(* CODESYS project JSON Utilities SL Example.project
   Title: JSON Utilities SL Example
   Author: CODESYS Development GmbH
   Company: CODESYS

Project tree, tasks and I/O mapping:
  Device : CODESYS Control for Raspberry Pi 64 SL, CODESYS, order no. 2302000009, version 4.18.0.0
    application JSONFindValueExample
      libraries: Standard, 3.5.18.0 (System); VisuDialogs, * (System); CAA FB Factory, * (CAA Technical Workgroup); JSON Utilities SL, 1.11.0.0 (CODESYS)
      task MainTask (cyclic, interval t#20ms, priority 1) calls PLC_PRG
      task VISU_TASK (cyclic, interval 100 ms, priority 31) calls VisuElems.Visu_Prg
      program PLC_PRG [CFC]
      visualisation Visualization
      image pool ImagePool
    application JSONFileExample
      libraries: Standard, 3.5.18.0 (System); VisuDialogs, * (System); CAA FB Factory, * (CAA Technical Workgroup); JSON Utilities SL, 1.11.0.0 (CODESYS)
      task MainTask (cyclic, interval t#20ms, priority 1) calls PLC_PRG
      task VISU_TASK (cyclic, interval 100 ms, priority 31) calls VisuElems.Visu_Prg
      program PLC_PRG [CFC]
      visualisation Visualization
      image pool ImagePool
    application JSONArrayExample
      libraries: Standard, 3.5.18.0 (System); VisuDialogs, * (System); CAA FB Factory, * (CAA Technical Workgroup); JSON Utilities SL, 1.11.0.0 (CODESYS)
      task MainTask (cyclic, interval t#20ms, priority 1) calls PLC_PRG
      task VISU_TASK (cyclic, interval 100 ms, priority 31) calls VisuElems.Visu_Prg
      program PLC_PRG [CFC]
      visualisation Visualization
      image pool ImagePool
    application JSONDataExample
      libraries: CAA FB Factory, * (CAA Technical Workgroup); JSON Utilities SL, 1.11.0.0 (CODESYS)
      task Task (cyclic, interval t#20ms, priority 1) calls PLC_PRG
      program PLC_PRG [ST]
    SoftMotion General Axis Pool
    GPIOs_A_B : GPIOs A/B, CODESYS, version 4.18.0.0
        unmapped channels: digital inputs (GPIO0..GPIO31), digital outputs (GPIO0..GPIO31)
    Onewire
    Camera device
      <Empty>
    SPI
    I²C
  text list GlobalTextList
  function block Element2StringArray [ST]
  5ce3da45-db07-42e7-a21c-a00fff4ed8f6|C:\Users\a.werner\Documents\background.jpg
  5ce3da45-db07-42e7-a21c-a00fff4ed8f6|C:\Users\a.werner\Documents\background.jpg
  5ce3da45-db07-42e7-a21c-a00fff4ed8f6|C:\Users\a.werner\Documents\background.jpg
*)

// Device/JSONFindValueExample/PLC_PRG
// This program loads the demo file 'test.json' and finds the value of the first key in the file. 
PROGRAM PLC_PRG
VAR
	sFileName : STRING(255) := 'res/test.json';	

	jsonDataFactory : JSON.JSONDataFactory;
	eDataFactoryError : FBF.ERROR; // Error code: 0: OK, 30103: no more memory 
	pJSONData : POINTER TO JSON.JSONData := jsonDataFactory.Create(eError => eDataFactoryError);

	JSONFileReader_0: JSON.JSONFileReader;
	xStart : BOOL;
	xFindValue : BOOL;
	wsKey : WSTRING := "Vorname";
	element : JSON.JSONElement;
	FindFirstValueByKey_0: JSON.FindFirstValueByKey;
	wsValue: WSTRING(JSON.GParams.g_diMaxStringSize);
END_VAR

// Load the example file 'c:\temp\test.json'
JSONFileReader_0(xExecute := xStart, sFileName := sFileName, jsonData := pJSONData^); // JSON.JSONFileReader
// Find a value by key
FindFirstValueByKey_0(xExecute := xFindValue, wsKey := wsKey, diStartIndex := 0, jsonData := pJSONData^); // JSON.FindFirstValueByKey
JSON.JSONElementToString(element := FindFirstValueByKey_0.jsonElement, wsResult := wsValue);

END_PROGRAM

// Device/JSONFileExample/PLC_PRG
// This program shows how to read and write JSON files.
PROGRAM PLC_PRG
VAR
	// JSON data container
	jsonDataFactory : JSON.JSONDataFactory; // Factory to create a JSONData function block. 
	eDataFactoryError : FBF.ERROR; // Error code: 0: OK, 30103: no more memory
	pJSONData : POINTER TO JSON.JSONData := jsonDataFactory.Create(eError => eDataFactoryError); // Result of Create is a pointer to JSONData
	
	// Reader
	JSONFileReader_0: JSON.JSONFileReader; 
	wsFilenameRead : STRING(255) := 'res/test.json';
	xReadFile : BOOL;
	
	// Writer
	JSONFileWriter_0: JSON.JSONFileWriter;
	wsFilenameWrite : STRING(255) := 'res/testWrite.json';
	xWriteFile : BOOL;
	
	// Helper array for visu
	awsData :  ARRAY[0..3, 0..500] OF WSTRING(JSON.GParams.g_diMaxStringSize);
	element2StringArray : Element2StringArray; // Function block to convert the sample data into an array of WSTRINGs (only for visualization)
END_VAR

// Convert the result into an array of WSTRINGs (only for visualization)
element2StringArray(xExecute := JSONFileReader_0.xDone, jsonData := pJSONData^, awsDataArray := awsData);
// Load the example file 'c:\temp\test.json'
JSONFileReader_0(xExecute := xReadFile, sFileName := wsFilenameRead, jsonData := pJSONData^); // JSON.JSONFileReader
// Write a JSON file
JSONFileWriter_0(
    xExecute := xWriteFile,
    sFileName := wsFilenameWrite,
    eEncoding := JSON.Encoding.UTF_8,
    jsonData := pJSONData^); // JSON.JSONFileWriter

END_PROGRAM

// Element2StringArray
// Helper function to convert the JSON elements to an array of WSTRINGs.
FUNCTION_BLOCK Element2StringArray
VAR_INPUT
	xExecute : BOOL; // Starts converting..
END_VAR
VAR_IN_OUT
	jsonData : JSON.JSONData;
	awsDataArray : ARRAY[0..3, 0..500] OF WSTRING(JSON.GParams.g_diMaxStringSize);
END_VAR
VAR
	diCounter : DINT;
	irow, icol : INT;
	element : JSON.JSONElement;
	j, i : INT;
END_VAR

IF xExecute = FALSE THEN
	RETURN;
END_IF
diCounter := 0;
irow := 0;
WHILE irow < 500 AND diCounter < JSON.GParams.g_diMaxElements DO
	jsonData.GetElementByIndex(diIndex := diCounter, jsonElement => element);
	IF element.eType = JSON.JSONType.NONE THEN
		FOR j := irow TO 500 DO
			FOR i := 0 TO 3 DO
				awsDataArray[i, j] := "";
			END_FOR	
		END_FOR
		RETURN;
	END_IF
	icol := 0;	
	
	// Index
	awsDataArray[icol, irow] := DINT_TO_WSTRING(element.diIndex);
	icol := icol + 1;
	
	// Parent Index
	awsDataArray[icol, irow] := DINT_TO_WSTRING(element.diParentIndex);
	icol := icol + 1;
	
	// Type
	IF element.eType = JSON.JSONType.BOOL_VALUE THEN
		awsDataArray[icol, irow] := "Bool";
	ELSIF element.eType = JSON.JSONType.LINT_VALUE THEN
		awsDataArray[icol, irow] := "LInt";
	ELSIF element.eType = JSON.JSONType.JSON_ARRAY THEN
		awsDataArray[icol, irow] := "Array";
	ELSIF element.eType = JSON.JSONType.JSON_OBJECT THEN
		awsDataArray[icol, irow] := "Object";
	ELSIF element.eType = JSON.JSONType.KEY THEN
		awsDataArray[icol, irow] := "Key";
	ELSIF element.eType = JSON.JSONType.NONE THEN
		awsDataArray[icol, irow] := "None";
	ELSIF element.eType = JSON.JSONType.NULL THEN
		awsDataArray[icol, irow] := "Null";
	ELSIF element.eType = JSON.JSONType.LREAL_VALUE THEN
		awsDataArray[icol, irow] := "LReal";
	ELSIF element.eType = JSON.JSONType.WSTRING_VALUE THEN
		awsDataArray[icol, irow] := "String";
	ELSE
		awsDataArray[icol, irow] := "Unknown";
	END_IF	
	icol := icol + 1;
	
	// Value
	IF element.eType = JSON.JSONType.BOOL_VALUE THEN
		awsDataArray[icol, irow] := BOOL_TO_WSTRING(element.value.xValue);
	ELSIF element.eType = JSON.JSONType.LINT_VALUE THEN
		awsDataArray[icol, irow] := LINT_TO_WSTRING(element.value.liValue);
	ELSIF element.eType = JSON.JSONType.KEY OR element.eType = JSON.JSONType.WSTRING_VALUE THEN
		awsDataArray[icol, irow] := element.value.wsValue;
	ELSIF element.eType = JSON.JSONType.LREAL_VALUE THEN
		awsDataArray[icol, irow] := LREAL_TO_WSTRING(element.value.lrValue);	
	ELSIF element.eType = JSON.JSONType.NULL THEN
		awsDataArray[icol, irow] := "Null";	
	ELSE
		awsDataArray[icol, irow] := "";	
	END_IF
	irow := irow + 1;
	diCounter := diCounter + 1;	
END_WHILE

END_FUNCTION_BLOCK

// Device/JSONArrayExample/PLC_PRG
// This program shows how to read and write JSON arrays.
PROGRAM PLC_PRG
VAR
	// JSON data container
	jsonDataFactory : JSON.JSONDataFactory; // Factory to create a JSONData function block. 
	eDataFactoryError : FBF.ERROR; // Error code: 0: OK, 30103: no more memory
	pJSONData : POINTER TO JSON.JSONData := jsonDataFactory.Create(eError => eDataFactoryError); // Result of Create is a pointer to JSONData
	
	// Reader
	JSONByteArrayReader_0: JSON.JSONByteArrayReader;	
	xRead : BOOL;
	// Demo data
	wsData : WSTRING(1024) := "{
  $0022Herausgeber$0022: $0022Xema$0022,
  $0022Nummer$0022: $00221234-5678-9012-3456$0022,
  $0022Deckung$0022: -0.444,
  $0022Waehrung$0022: $0022EURO$0022,
  $0022Inhaber$0022: 
  {
    $0022Name$0022: $0022Mustermann$0022,
    $0022Vorname$0022: $0022Max$0022,
    $0022maennlich$0022: true,
    $0022Hobbys$0022: [ $0022Reiten$0022, $0022Golfen$0022, $0022Lesen$0022 ],
    $0022Alter$0022: 42,
    $0022Kinder$0022: [],
    $0022Partner$0022: null
  }
}";
	
	// Writer
	JSONByteArrayWriter_0: JSON.JSONByteArrayWriter;
	wsWriteData : WSTRING(1024) := ""; // The result of the Writer
	xWrite : BOOL;
	
	// Helper array for visu
	awsData :  ARRAY[0..3, 0..500] OF WSTRING(JSON.GParams.g_diMaxStringSize);	
	element2StringArray : Element2StringArray; // Function block to convert the sample data into an array of WSTRINGs (only for visualization)
END_VAR

// Read JSON data from WSTRING
JSONByteArrayReader_0(xExecute := xRead, pwData := ADR(wsData), jsonData := pJSONData^); // JSON.JSONByteArrayReader
// Convert the result into an array of WSTRINGs (only for visualization)
element2StringArray(xExecute := JSONByteArrayReader_0.xDone, jsonData := pJSONData^, awsDataArray := awsData);
// Read JSON data to WSTRING
JSONByteArrayWriter_0(
    xExecute := xWrite,
    pwData := ADR(wsWriteData),
    udiSize := SIZEOF(wsWriteData),
    jsonData := pJSONData^); // JSON.JSONByteArrayWriter

END_PROGRAM

// Device/JSONDataExample/PLC_PRG
// This program shows how to build a JSON data string.
PROGRAM PLC_PRG
VAR
	factory : JSON.JSONDataFactory;
	eDataFactoryError : FBF.ERROR; // Error code: 0: OK, 30103: no more memory	
	pJsonData : POINTER TO JSON.JSONData := factory.Create(eError => eDataFactoryError);
	jsonArrayWriter : JSON.JSONByteArrayWriter; 
	diCounter : DINT;
	diMemory : DINT;
	wsJsonData : WSTRING(1000); 
	wsValue : WSTRING;
	xStart : BOOL := TRUE;
	iExample : INT := 1; // Default example 1
	fb_JBuilder : JSON.JSONBuilder;
	xValue : BOOL := TRUE;
	iValue : INT := 42;
	lrValue : LREAL := -0.444;
	wsArrValue : ARRAY [0..2] OF WSTRING := ["Reiten", "Golfen", "Lesen"];
END_VAR

IF xStart = TRUE AND pJsonData <> 0 THEN
	IF iExample = 1 THEN
		diCounter := 0;
		// Index of the root object is -1.
		pJsonData^.SetObject(diIndex := diCounter, diParentIndex := -1);
		diCounter := diCounter + 1;
		// The parent index of the key is the index of parent object.
		pJsonData^.SetKey(wsKey := "Key1", diParentIndex := 0, diIndex := diCounter);
		diCounter := diCounter + 1;
		// The parent index of the value is the index of corresponding key.
		pJsonData^.SetString(wsValue := "Value1", diIndex := diCounter, diParentIndex := diCounter - 1);
		
		diCounter := diCounter + 1;
		pJsonData^.SetKey(wsKey := "Key2", diParentIndex := 0, diIndex := diCounter);
		diCounter := diCounter + 1;
		pJsonData^.SetLInt(liValue := 77, diIndex := diCounter, diParentIndex := diCounter - 1);
		
		diCounter := diCounter + 1;
		pJsonData^.SetKey(wsKey := "Key3", diParentIndex := 0, diIndex := diCounter);
		diCounter := diCounter + 1;
		pJsonData^.SetBool(bValue := FALSE, diIndex := diCounter, diParentIndex := diCounter - 1);	
	END_IF
	// This example recreates the test.json file
	IF iExample = 2 THEN
		// Initialize fb and set root object
		fb_JBuilder(pJsonData := pJsonData, diRootObj => diCounter);
		wsValue := "Xema";
		// JSON:    "Herausgeber": "Xema", 
		fb_JBuilder.SetKeyWithValue("Herausgeber", wsValue, diParentIndex := diCounter);
		wsValue := "1234-5678-9012-3456";
		// JSON:   "Nummer": "1234-5678-9012-3456", 
		fb_JBuilder.SetKeyWithValue("Nummer", wsValue, diCounter);
		// JSON:   "Deckung": -4.44e-1, 
		fb_JBuilder.SetKeyWithValue("Deckung", lrValue, diCounter);
		wsValue := "EURO";
		// JSON:    "Waehrung": "EURO", 
		fb_JBuilder.SetKeyWithValue("Waehrung", wsValue, diCounter);
		// Set key with object, and override diParent. JSON:    "Inhaber": {
		diCounter := fb_JBuilder.SetKeyWithObject("Inhaber", diCounter);
		wsValue := "\ $"Mustermann\$"";
		// JSON:       "Name": "\ \"Mustermann\\"", 
		fb_JBuilder.SetKeyWithValue("Name", wsValue, diCounter);
		wsValue := "Max";
		// JSON:       "Vorname": "Max", 
		fb_JBuilder.SetKeyWithValue("Vorname", wsValue, diCounter);
		// JSON:       "maennlich": true, 
		fb_JBuilder.SetKeyWithValue("maennlich", xValue, diCounter);
		// Save parent to use after it after the array again
		diMemory := diCounter;
		// JSON:       "Hobbys": 
		diCounter := fb_JBuilder.SetKeyWithArray("Hobbys", diCounter);
		// JSON:         ["Reiten", "Golfen", "Lesen"],
		fb_JBuilder.SetValue(wsArrValue[0], diCounter);
		fb_JBuilder.SetValue(wsArrValue[1], diCounter);
		fb_JBuilder.SetValue(wsArrValue[2], diCounter);
		// Use saved parent. JSON:       "Alter": 42, 
		fb_JBuilder.SetKeyWithValue("Alter", iValue, diMemory);
		// JSON:       "Kinder": 
		// JSON:         [],
		fb_JBuilder.SetKeyWithArray("Kinder", diMemory);
		// JSON:       "Partner": null
		fb_JBuilder.SetKeyWithValueNull("Partner", diMemory);
	END_IF
	xStart := FALSE;
END_IF

// Generate the JSON String. The value will be written to the variable wsJsonData.
jsonArrayWriter(xExecute := TRUE, pwData := ADR(wsJsonData), udiSize := SIZEOF(wsJsonData), jsonData := pJsonData^);

END_PROGRAM

// Device/JSONFindValueExample/Visualization
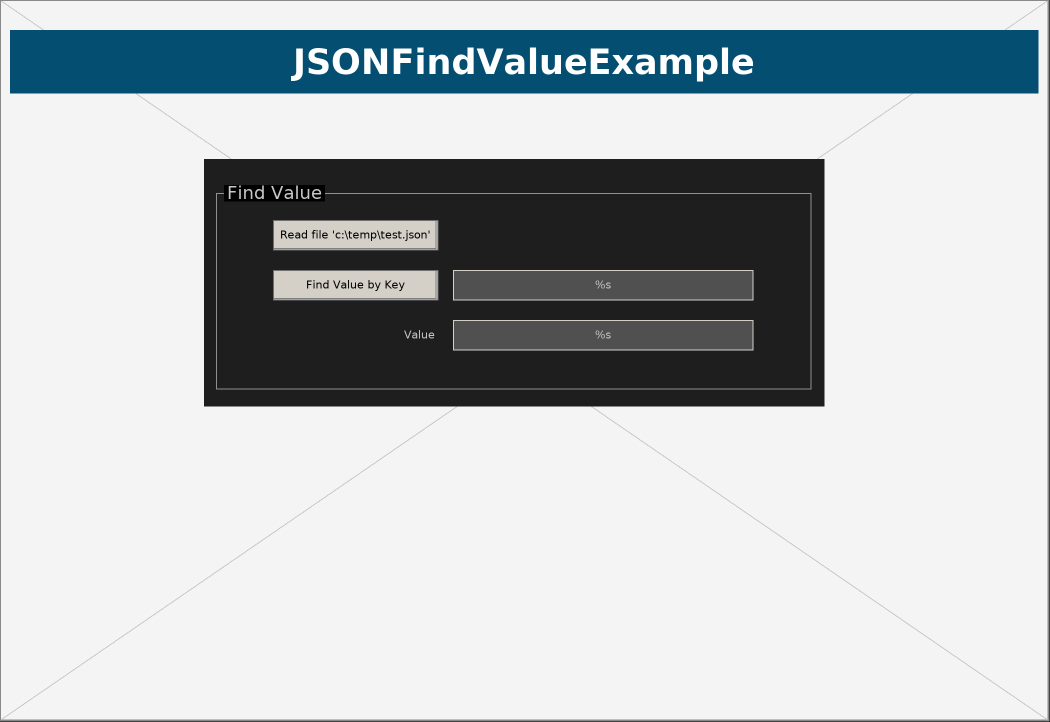
VISUALIZATION Visualization  // 1050x722
    Image (0,0 1048x720), image: ImagePool.Background
    Rectangle (204,159 620x247)
    GroupBox (216,185 595x204), "Find Value"
        Group (57,35 480x130)
            Button (0,0 165x30), "Read file 'c:\temp\test.json'"
                tap PLC_PRG.xStart
            Button (0,50 165x30), "Find Value by Key"
                tap PLC_PRG.xFindValue
            Textfield (180,50 300x30), "%s", text variable: PLC_PRG.wsKey
                OnMouseClick: write the text variable via Default
            Textfield (180,100 300x30), "%s", text variable: PLC_PRG.wsValue
            Label (0,100 165x30), "Value"
    Rectangle (10,30 1028x63), "JSONFindValueExample"
END_VISUALIZATION

// Device/JSONFileExample/Visualization
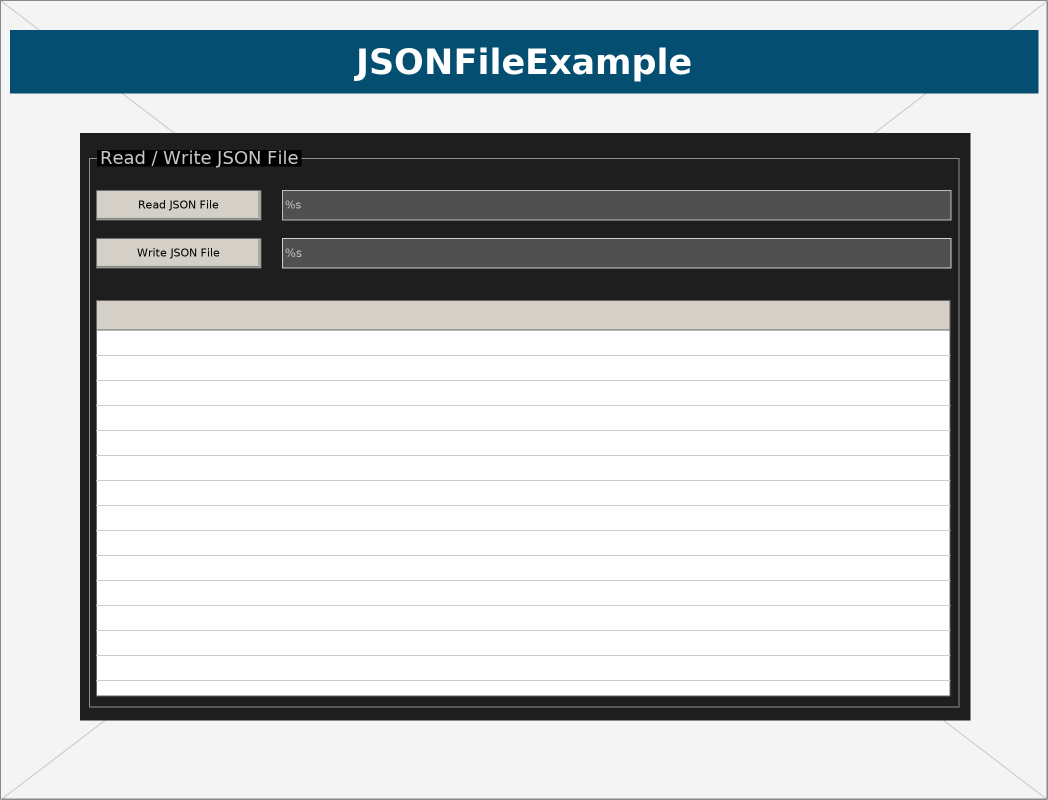
VISUALIZATION Visualization  // 1048x800
    Image (0,0 1048x800), image: ImagePool.background
    Rectangle (80,133 890x587)
    GroupBox (89,150 870x557), "Read / Write JSON File"
        Group (7,40 855x78)
            Button (0,0 165x30), "Read JSON File"
                tap PLC_PRG.xReadFile
            Textfield (186,0 669x30), "%s", text variable: PLC_PRG.wsFilenameRead
                OnMouseClick: write the text variable via Default
            Button (0,48 165x30), "Write JSON File"
                tap PLC_PRG.xWriteFile
            Textfield (186,48 669x30), "%s", text variable: PLC_PRG.wsFilenameWrite
                OnMouseClick: write the text variable via Default
        Table (7,150 854x396), data array: PLC_PRG.awsData
            p3854506369: PLC_PRG.awsData[0,INDEX]
            p1892666644: PLC_PRG.awsData[1,INDEX]
            p338671338: PLC_PRG.awsData[2,INDEX]
            p2170511999: PLC_PRG.awsData[3,INDEX]
            p2232123230: Index
            p511219082: Parent Index
            p1755163831: Type
            p4092479075: Value
    Rectangle (10,30 1028x63), "JSONFileExample"
END_VISUALIZATION

// Device/JSONArrayExample/Visualization
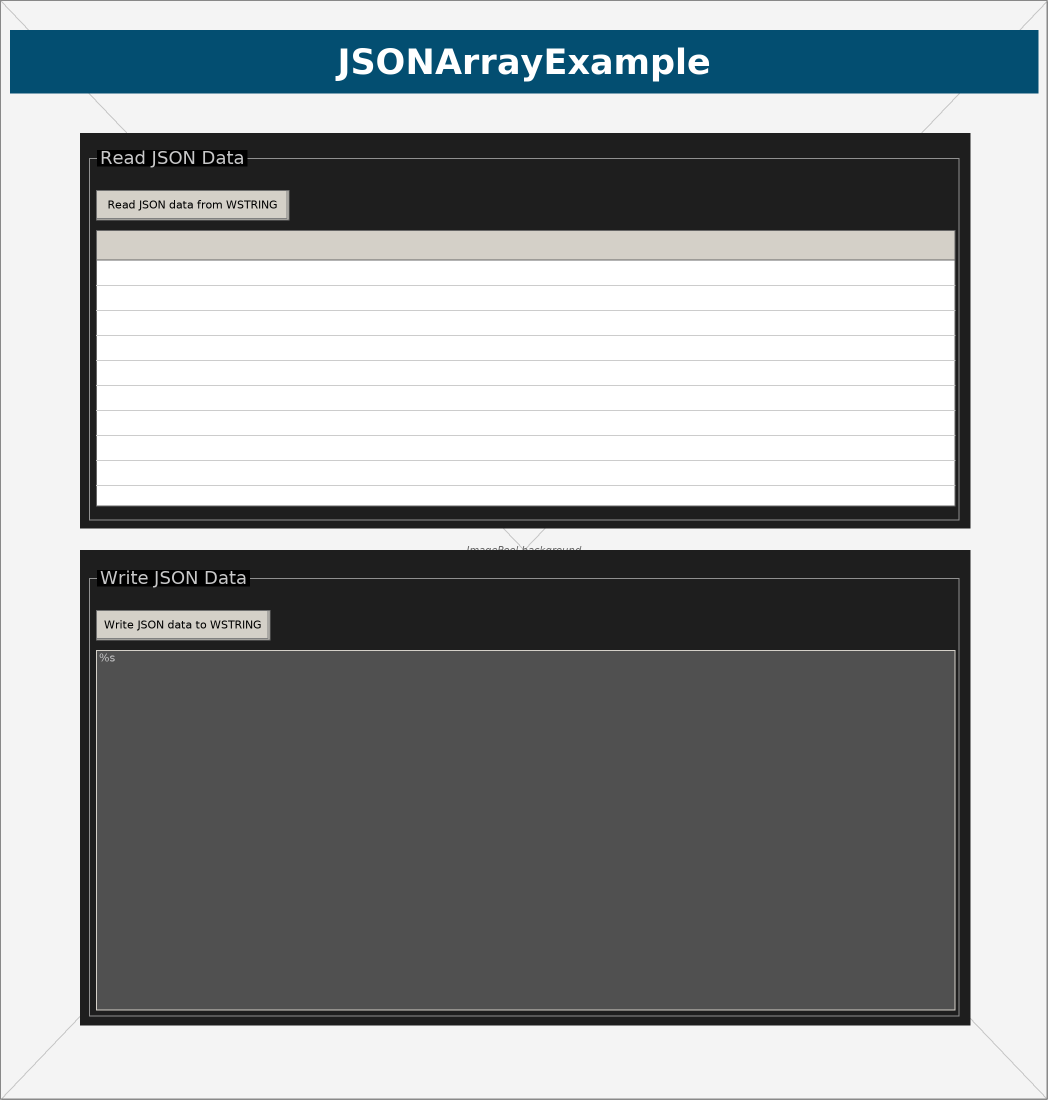
VISUALIZATION Visualization  // 1048x1100
    Image (0,0 1048x1100), image: ImagePool.background
    Rectangle (80,550 890x475)
    Rectangle (80,133 890x395)
    GroupBox (89,570 870x446), "Write JSON Data"
        Button (7,40 174x30), "Write JSON data to WSTRING"
            tap PLC_PRG.xWrite
        Textfield (7,80 859x360), "%s", text variable: PLC_PRG.wsWriteData
    GroupBox (89,150 870x370), "Read JSON Data"
        Button (7,40 193x30), "Read JSON data from WSTRING"
            tap PLC_PRG.xRead
        Table (7,80 859x276), data array: PLC_PRG.awsData
            p3854506369: PLC_PRG.awsData[0,INDEX]
            p1892666644: PLC_PRG.awsData[1,INDEX]
            p338671338: PLC_PRG.awsData[2,INDEX]
            p2170511999: PLC_PRG.awsData[3,INDEX]
            p2232123230: Index
            p511219082: Parent Index
            p1755163831: Type
            p4092479075: Value
    Rectangle (10,30 1028x63), "JSONArrayExample"
END_VISUALIZATION
